   "80_From_HMI_MAN_DQ_139_4" : Bool = PLC "80_From_HMI".MAN_DQ_139_4, 1 s
   "80_From_HMI_MAN_DQ_139_5" : Bool = PLC "80_From_HMI".MAN_DQ_139_5, 1 s
   "80_From_HMI_MAN_DQ_139_6" : Bool = PLC "80_From_HMI".MAN_DQ_139_6, 1 s
   "80_From_HMI_MAN_DQ_139_7" : Bool = PLC "80_From_HMI".MAN_DQ_139_7, 1 s
   "80_From_HMI_P301_PRSNT" : Bool = PLC "80_From_HMI".P301_PRSNT, 1 s
   "80_From_HMI_P305_PRSNT" : Bool = PLC "80_From_HMI".P305_PRSNT, 1 s
   "80_From_HMI_PIT 316 delay" : Time = PLC "80_From_HMI"."PIT 316 delay", 1 s
   "80_From_HMI_PIT 359 delay" : Time = PLC "80_From_HMI"."PIT 359 delay", 1 s
   "80_From_HMI_Post Purge Time" : Time = PLC "80_From_HMI"."Post Purge Time", 1 s
   "80_From_HMI_Request_Auto" : Bool = PLC "80_From_HMI".Request_Auto, 1 s
   "80_From_HMI_Request_Manual" : Bool = PLC "80_From_HMI".Request_Manual, 1 s
   "80_From_HMI_Reset CV203 PID" : Bool = PLC "80_From_HMI"."Reset CV203 PID", 1 s
   "80_From_HMI_Reset_Alarms" : Bool = PLC "80_From_HMI".Reset_Alarms, 1 s
   "80_From_HMI_RST_AUT_SEQ" : Bool = PLC "80_From_HMI".RST_AUT_SEQ, 1 s
   "80_From_HMI_RST_LOCKOUT" : Bool = PLC "80_From_HMI".RST_LOCKOUT, 1 s
   "80_From_HMI_RUN_BTCS" : Bool = PLC "80_From_HMI".RUN_BTCS, 1 s
   "80_From_HMI_RUN_BWTS" : Bool = PLC "80_From_HMI".RUN_BWTS, 1 s
   "80_From_HMI_SAL_CNFRM" : Bool = PLC "80_From_HMI".SAL_CNFRM, 1 s
   "80_From_HMI_SAL_VALUE" : Real = PLC "80_From_HMI".SAL_VALUE, 1 s
   "80_From_HMI_Test Tank Request" : Bool = PLC "80_From_HMI"."Test Tank Request", 1 s
   "80_From_HMI_TIMER RST Supres" : Bool = PLC "80_From_HMI"."TIMER RST Supres", 1 s
   "82_To_HMI_CA Blower Reset Hours" : Bool = PLC "82_To_HMI"."CA Blower Reset Hours", 1 s
   "82_To_HMI_CA Blower Run Seconds" : Int = PLC "82_To_HMI"."CA Blower Run Seconds", 1 s
   "82_To_HMI_CA Blower Service Due" : Bool = PLC "82_To_HMI"."CA Blower Service Due", 1 s
   "82_To_HMI_CA Blower Total Run Hours" : Int = PLC "82_To_HMI"."CA Blower Total Run Hours", 1 s
   "82_To_HMI_CRNT_MODE" : Int = PLC "82_To_HMI".CRNT_MODE_IGG, 1 s
   "82_To_HMI_CRNT_MODE_GCU" : Int = PLC "82_To_HMI".CRNT_MODE_GCU, 1 s
   "82_To_HMI_E500A Fuel Pump Reset Hours" : Bool = PLC "82_To_HMI"."E500A Fuel Pump Reset Hours", 1 s
   "82_To_HMI_E500A Fuel Pump Run Hours" : Int = PLC "82_To_HMI"."E500A Fuel Pump Run Hours", 1 s
   "82_To_HMI_E500A Fuel Pump Run Minutes" : Int = PLC "82_To_HMI"."E500A Fuel Pump Run Minutes", 1 s
   "82_To_HMI_E500A Fuel Pump Run Seconds" : Int = PLC "82_To_HMI"."E500A Fuel Pump Run Seconds", 1 s
   "82_To_HMI_E500A Fuel Pump Service Due" : Bool = PLC "82_To_HMI"."E500A Fuel Pump Service Due", 1 s
   "82_To_HMI_E500A Fuel Pump Service Time Hours" : Int = PLC "82_To_HMI"."E500A Fuel Pump Service Time Hours", 1 s
   "82_To_HMI_E500A Fuel Pump Total Run Hours" : Int = PLC "82_To_HMI"."E500A Fuel Pump Total Run Hours", 1 s
   "82_To_HMI_E500B Fuel Pump Reset Hours" : Bool = PLC "82_To_HMI"."E500B Fuel Pump Reset Hours", 1 s
   "82_To_HMI_E500B Fuel Pump Run Minutes" : Int = PLC "82_To_HMI"."E500B Fuel Pump Run Minutes", 1 s
   "82_To_HMI_E500B Fuel Pump Run Seconds" : Int = PLC "82_To_HMI"."E500B Fuel Pump Run Seconds", 1 s
   "82_To_HMI_E500B Fuel Pump Service Due" : Bool = PLC "82_To_HMI"."E500B Fuel Pump Service Due", 1 s
   "82_To_HMI_E500B Fuel Pump Service Time Hours" : Int = PLC "82_To_HMI"."E500B Fuel Pump Service Time Hours", 1 s
   "82_To_HMI_E500B Fuel Pump Total Run Hours" : Int = PLC "82_To_HMI"."E500B Fuel Pump Total Run Hours", 1 s
   "82_To_HMI_E-STOP LATCHED" : Bool = PLC "82_To_HMI"."E-STOP LATCHED", 1 s
   "82_To_HMI_I&A Compressor Reset Hours" : Bool = PLC "82_To_HMI"."I&A Compressor Reset Hours", 1 s
   "82_To_HMI_I&A Compressor Service Due" : Bool = PLC "82_To_HMI"."I&A Compressor Service Due", 1 s
   "82_To_HMI_I&A Compressor Total Run Hours" : Int = PLC "82_To_HMI"."I&A Compressor Total Run Hours", 1 s
   "82_To_HMI_P301 CSW Pump Reset Hours" : Bool = PLC "82_To_HMI"."P301 CSW Pump Reset Hours", 1 s
   "82_To_HMI_P301 CSW Pump Run Days" : Int = PLC "82_To_HMI"."P301 CSW Pump Run Days", 1 s
   "82_To_HMI_P301 CSW Pump Run Hours" : Int = PLC "82_To_HMI"."P301 CSW Pump Run Hours", 1 s
   "82_To_HMI_P301 CSW Pump Run Minutes" : Int = PLC "82_To_HMI"."P301 CSW Pump Run Minutes", 1 s
   "82_To_HMI_P301 CSW Pump Run Seconds" : Int = PLC "82_To_HMI"."P301 CSW Pump Run Seconds", 1 s
   "82_To_HMI_P301 CSW Pump Service Due" : Bool = PLC "82_To_HMI"."P301 CSW Pump Service Due", 1 s
   "82_To_HMI_P301 CSW Pump Service Time Hours" : Int = PLC "82_To_HMI"."P301 CSW Pump Service Time Hours", 1 s
   "82_To_HMI_P301 CSW Pump Total Run Hours" : Int = PLC "82_To_HMI"."P301 CSW Pump Total Run Hours", 1 s
   "82_To_HMI_P305 FW Pump Reset Hours" : Bool = PLC "82_To_HMI"."P305 FW Pump Reset Hours", 1 s
   "82_To_HMI_P305 FW Pump Run Days" : Int = PLC "82_To_HMI"."P305 FW Pump Run Days", 1 s
   "82_To_HMI_P305 FW Pump Run Hours" : Int = PLC "82_To_HMI"."P305 FW Pump Run Hours", 1 s
   "84_Setpoints_D_ON" : Bool = PLC "84_Setpoints".D_ON, 1 s
   "84_Setpoints_Derive Time" : Time = PLC "84_Setpoints"."Derive Time", 1 s
   "84_Setpoints_E400_PT002_High" : Real = PLC "84_Setpoints".E400_PT002_High, 1 s
   "84_Setpoints_E400_PT002_HighHigh" : Real = PLC "84_Setpoints".E400_PT002_HighHigh, 1 s
   "84_Setpoints_E400_TT002_High" : Real = PLC "84_Setpoints".E400_TT002_High, 1 s
   "84_Setpoints_E400_TT002_HighHigh" : Real = PLC "84_Setpoints".E400_TT002_HighHigh, 1 s
   "84_Setpoints_Gain" : Real = PLC "84_Setpoints".Gain, 1 s
   "84_Setpoints_I_ON" : Bool = PLC "84_Setpoints".I_ON, 1 s
   "84_Setpoints_Integration Time" : Time = PLC "84_Setpoints"."Integration Time", 1 s
   "84_Setpoints_LIT304_InitialFill_High" : Real = PLC "84_Setpoints".LIT304_InitialFill_High, 1 s
   "84_Setpoints_LIT304_InitialFill_HighHigh" : Real = PLC "84_Setpoints".LIT304_InitialFill_HighHigh, 1 s
   "84_Setpoints_LIT304_InitialFill_Low" : Real = PLC "84_Setpoints".LIT304_InitialFill_Low, 1 s
   "84_Setpoints_LIT304_InitialFill_LowLow" : Real = PLC "84_Setpoints".LIT304_InitialFill_LowLow, 1 s
   "84_Setpoints_LIT304_InitialFill_Target" : Real = PLC "84_Setpoints".LIT304_InitialFill_Target, 1 s
   "84_Setpoints_LIT304_InitialFill_Target_Low" : Real = PLC "84_Setpoints".LIT304_InitialFill_Target_Low, 1 s
   "84_Setpoints_LIT304_Refill_High" : Real = PLC "84_Setpoints".LIT304_Refill_High, 1 s
   "84_Setpoints_LIT304_Refill_HighHigh" : Real = PLC "84_Setpoints".LIT304_Refill_HighHigh, 1 s
   "84_Setpoints_LIT304_Refill_Low" : Real = PLC "84_Setpoints".LIT304_Refill_Low, 1 s
   "84_Setpoints_LIT304_Refill_LowLow" : Real = PLC "84_Setpoints".LIT304_Refill_LowLow, 1 s
   "84_Setpoints_LIT304_Refill_Target" : Real = PLC "84_Setpoints".LIT304_Refill_Target, 1 s
   "84_Setpoints_LIT304_Refill_Target_Low" : Real = PLC "84_Setpoints".LIT304_Refill_Target_Low, 1 s
   "84_Setpoints_Max Opening" : Real = PLC "84_Setpoints"."Max Opening", 1 s
   "84_Setpoints_Min Opening" : Real = PLC "84_Setpoints"."Min Opening", 1 s
   "84_Setpoints_P_ON" : Bool = PLC "84_Setpoints".P_ON, 1 s
   "84_Setpoints_PIT113_Burner_Target" : Real = PLC "84_Setpoints".PIT113_Burner_Target, 1 s
   "84_Setpoints_PIT204_High" : Real = PLC "84_Setpoints".PIT204_High, 1 s
   "84_Setpoints_PIT204_High(1)" : Real = PLC "84_Setpoints".PIT204_High, 1 s
   "84_Setpoints_PIT204_HighHigh" : Real = PLC "84_Setpoints".PIT204_HighHigh, 1 s
   "84_Setpoints_PIT204_HighHigh(1)" : Real = PLC "84_Setpoints".PIT204_HighHigh, 1 s
   "84_Setpoints_PIT204_Low" : Real = PLC "84_Setpoints".PIT204_Low, 1 s
   "84_Setpoints_PIT204_Low(1)" : Real = PLC "84_Setpoints".PIT204_Low, 1 s
   "84_Setpoints_PIT204_LowLow" : Real = PLC "84_Setpoints".PIT204_LowLow, 1 s
   "84_Setpoints_PIT204_LowLow(1)" : Real = PLC "84_Setpoints".PIT204_LowLow, 1 s
   "84_Setpoints_PIT348_High" : Real = PLC "84_Setpoints".PIT348_High, 1 s
   "84_Setpoints_PIT348_HighHigh" : Real = PLC "84_Setpoints".PIT348_HighHigh, 1 s
   "84_Setpoints_PIT348_Low" : Real = PLC "84_Setpoints".PIT348_Low, 1 s
   "84_Setpoints_PIT348_LowLow" : Real = PLC "84_Setpoints".PIT348_LowLow, 1 s
   "84_Setpoints_PIT353_InitialFill_High" : Real = PLC "84_Setpoints".PIT353_InitialFill_High, 1 s
   "84_Setpoints_PIT353_InitialFill_HighHigh" : Real = PLC "84_Setpoints".PIT353_InitialFill_HighHigh, 1 s
   "84_Setpoints_PIT353_InitialFill_Low" : Real = PLC "84_Setpoints".PIT353_InitialFill_Low, 1 s
   "84_Setpoints_PIT353_InitialFill_LowLow" : Real = PLC "84_Setpoints".PIT353_InitialFill_LowLow, 1 s
   "84_Setpoints_PIT353_Refill_High" : Real = PLC "84_Setpoints".PIT353_Refill_High, 1 s
   "84_Setpoints_PIT353_Refill_HighHigh" : Real = PLC "84_Setpoints".PIT353_Refill_HighHigh, 1 s
   "84_Setpoints_PIT353_Refill_Low" : Real = PLC "84_Setpoints".PIT353_Refill_Low, 1 s
   "84_Setpoints_PIT353_Refill_LowLow" : Real = PLC "84_Setpoints".PIT353_Refill_LowLow, 1 s
   "84_Setpoints_PIT358_InitialFill_High" : Real = PLC "84_Setpoints".PIT358_InitialFill_High, 1 s
   "84_Setpoints_PIT358_InitialFill_HighHigh" : Real = PLC "84_Setpoints".PIT358_InitialFill_HighHigh, 1 s
   "84_Setpoints_PIT358_InitialFill_Low" : Real = PLC "84_Setpoints".PIT358_InitialFill_Low, 1 s
   "84_Setpoints_PIT358_InitialFill_LowLow" : Real = PLC "84_Setpoints".PIT358_InitialFill_LowLow, 1 s
   "84_Setpoints_PIT358_Refill_High" : Real = PLC "84_Setpoints".PIT358_Refill_High, 1 s
   "84_Setpoints_PIT358_Refill_HighHigh" : Real = PLC "84_Setpoints".PIT358_Refill_HighHigh, 1 s
   "84_Setpoints_PIT358_Refill_Low" : Real = PLC "84_Setpoints".PIT358_Refill_Low, 1 s
   "84_Setpoints_PIT358_Refill_LowLow" : Real = PLC "84_Setpoints".PIT358_Refill_LowLow, 1 s
   "84_Setpoints_PIT416_High" : Real = PLC "84_Setpoints".PIT416_High, 1 s
   "84_Setpoints_PIT416_HighHigh" : Real = PLC "84_Setpoints".PIT416_HighHigh, 1 s
   "84_Setpoints_PIT416_Low" : Real = PLC "84_Setpoints".PIT416_Low, 1 s
   "84_Setpoints_PIT416_LowLow" : Real = PLC "84_Setpoints".PIT416_LowLow, 1 s
   "84_Setpoints_PIT416_Target" : Real = PLC "84_Setpoints".PIT416_Target, 1 s
   "84_Setpoints_TIT406_High" : Real = PLC "84_Setpoints".TIT406_High, 1 s
   "84_Setpoints_TIT406_HighHigh" : Real = PLC "84_Setpoints".TIT406_HighHigh, 1 s
   "84_Setpoints_TIT408_High" : Real = PLC "84_Setpoints".TIT408_High, 1 s
   "84_Setpoints_TIT408_HighHigh" : Real = PLC "84_Setpoints".TIT408_HighHigh, 1 s
   "86_Times_CV341_CLSD_DLY" : Time = PLC "86_Times".CV341_CLSD_DLY, 1 s
   "86_Times_CV341_MAX_TRVL_TIME" : Time = PLC "86_Times".CV341_MAX_TRVL_TIME, 1 s
   "86_Times_CV341_OPND_DLY" : Time = PLC "86_Times".CV341_OPND_DLY, 1 s
   "86_Times_CV358_CLSD_DLY" : Time = PLC "86_Times".CV358_CLSD_DLY, 1 s
   "86_Times_CV358_MAX_TRVL_TIME" : Time = PLC "86_Times".CV358_MAX_TRVL_TIME, 1 s
   "86_Times_CV401_CLSD_DLY" : Time = PLC "86_Times".CV401_CLSD_DLY, 1 s
   "86_Times_CV401_OPND_DLY" : Time = PLC "86_Times".CV401_OPND_DLY, 1 s
   "86_Times_CV405_OPND_DLY" : Time = PLC "86_Times".CV405_OPND_DLY, 1 s
   "86_Times_CV406_CLSD_DLY" : Time = PLC "86_Times".CV406_CLSD_DLY, 1 s
   "86_Times_CV406_MAX_TRVL_TIME" : Time = PLC "86_Times".CV406_MAX_TRVL_TIME, 1 s
   "86_Times_CV407_MAX_TRVL_TIME" : Time = PLC "86_Times".CV407_MAX_TRVL_TIME, 1 s
   "86_Times_CV409_MAX_TRVL_TIME" : Time = PLC "86_Times".CV409_MAX_TRVL_TIME, 1 s
   "86_Times_CV411_MAX_TRVL_TIME" : Time = PLC "86_Times".CV411_MAX_TRVL_TIME, 1 s
   "86_Times_CV441_CLSD_DLY" : Time = PLC "86_Times".CV441_CLSD_DLY, 1 s
   "86_Times_CV441_MAX_TRVL_TIME" : Time = PLC "86_Times".CV441_MAX_TRVL_TIME, 1 s
   "86_Times_CV441_OPND_DLY" : Time = PLC "86_Times".CV441_OPND_DLY, 1 s
   "86_Times_E400_RNG_DLY" : Time = PLC "86_Times".E400_RNG_DLY, 1 s
   "86_Times_E400_STOP_TIME" : Time = PLC "86_Times".E400_STOP_TIME, 1 s
   "86_Times_E400_STRTD_DLY" : Time = PLC "86_Times".E400_STRTD_DLY, 1 s
   "86_Times_GCU_FLUSH_TIME" : Time = PLC "86_Times".GCU_FLUSH_TIME, 1 s
   "86_Times_GCU_TNK_DRN_MAX_TIME" : Time = PLC "86_Times".GCU_TNK_DRN_MAX_TIME, 1 s
   "86_Times_GCU_TNK_FILL_MAX_TIME" : Time = PLC "86_Times".GCU_TNK_FILL_MAX_TIME, 1 s
   "86_Times_LIT304 Delay" : Time = PLC "86_Times"."LIT304 Delay", 1 s
   "86_Times_P301_START_DLY" : Time = PLC "86_Times".P301_START_DLY, 1 s
   "86_Times_P303_STOP_TIME" : Time = PLC "86_Times".P303_STOP_TIME, 1 s
   "86_Times_P303_STPD_DLY" : Time = PLC "86_Times".P303_STPD_DLY, 1 s
   "86_Times_P303_STRTD_DLY" : Time = PLC "86_Times".P303_STRTD_DLY, 1 s
   "86_Times_P304_STPD_DLY" : Time = PLC "86_Times".P304_STPD_DLY, 1 s
   "86_Times_P304_STRTD_DLY" : Time = PLC "86_Times".P304_STRTD_DLY, 1 s
   "86_Times_P305_STPD_DLY" : Time = PLC "86_Times".P305_STPD_DLY, 1 s
   "86_Times_P305_STRTD_DLY" : Time = PLC "86_Times".P305_STRTD_DLY, 1 s
   "86_Times_PIT353 Delay" : Time = PLC "86_Times"."PIT353 Delay", 1 s
   "86_Times_PIT402 Alarm Delay" : Time = PLC "86_Times"."PIT402 Alarm Delay", 1 s
   "86_Times_PIT402_Ramp_Seconds" : Int = PLC "86_Times".PIT402_Ramp_Seconds, 1 s
   "86_Times_PIT416 Delay" : Time = PLC "86_Times"."PIT416 Delay", 1 s
   "86_Times_PIT416_TRGT_RMP_TIME" : Real = PLC "86_Times".PIT416_TRGT_RMP_TIME, 1 s
   "86_Times_POST_FLUSH_DLY" : Time = PLC "86_Times".POST_FLUSH_DLY, 1 s
   "86_Times_PRE_CV441_OPN_DLY" : Time = PLC "86_Times".PRE_CV441_OPN_DLY, 1 s
   "86_Times_PRE_GCU_TNK_FILL_DLY" : Time = PLC "86_Times".PRE_GCU_TNK_FILL_DLY, 1 s
   "86_Times_STEP_MAX_TIME_STP_001" : Time = PLC "86_Times".STEP_MAX_TIME_STP_001, 1 s
   "86_Times_STEP_MAX_TIME_STP_005" : Time = PLC "86_Times".STEP_MAX_TIME_STP_005, 1 s
   "86_Times_STEP_MAX_TIME_STP_010" : Time = PLC "86_Times".STEP_MAX_TIME_STP_010, 1 s
   "86_Times_STEP_MAX_TIME_STP_020" : Time = PLC "86_Times".STEP_MAX_TIME_STP_020, 1 s
   "86_Times_STEP_MAX_TIME_STP_030" : Time = PLC "86_Times".STEP_MAX_TIME_STP_030, 1 s
   "86_Times_STEP_MAX_TIME_STP_040" : Time = PLC "86_Times".STEP_MAX_TIME_STP_040, 1 s
   "86_Times_STEP_MAX_TIME_STP_050" : Time = PLC "86_Times".STEP_MAX_TIME_STP_050, 1 s
   "86_Times_STEP_MAX_TIME_STP_060" : Time = PLC "86_Times".STEP_MAX_TIME_STP_060, 1 s
   "86_Times_STEP_MAX_TIME_STP_070" : Time = PLC "86_Times".STEP_MAX_TIME_STP_070, 1 s
   "86_Times_STEP_MAX_TIME_STP_080" : Time = PLC "86_Times".STEP_MAX_TIME_STP_080, 1 s
   "86_Times_STEP_MAX_TIME_STP_090" : Time = PLC "86_Times".STEP_MAX_TIME_STP_090, 1 s
   "86_Times_STEP_MAX_TIME_STP_100" : Time = PLC "86_Times".STEP_MAX_TIME_STP_100, 1 s
   "86_Times_STEP_MAX_TIME_STP_110" : Time = PLC "86_Times".STEP_MAX_TIME_STP_110, 1 s
   "86_Times_STEP_MAX_TIME_STP_120" : Time = PLC "86_Times".STEP_MAX_TIME_STP_120, 1 s
   "86_Times_STEP_MAX_TIME_STP_130" : Time = PLC "86_Times".STEP_MAX_TIME_STP_130, 1 s
   "86_Times_STEP_MAX_TIME_STP_140" : Time = PLC "86_Times".STEP_MAX_TIME_STP_140, 1 s
   "86_Times_STEP_MAX_TIME_STP_150" : Time = PLC "86_Times".STEP_MAX_TIME_STP_150, 1 s
   "86_Times_STEP_MAX_TIME_STP_160" : Time = PLC "86_Times".STEP_MAX_TIME_STP_160, 1 s
   "86_Times_STEP_MAX_TIME_STP_170" : Time = PLC "86_Times".STEP_MAX_TIME_STP_170, 1 s
   "86_Times_STEP_MAX_TIME_STP_180" : Time = PLC "86_Times".STEP_MAX_TIME_STP_180, 1 s
   "86_Times_STEP_MAX_TIME_STP_190" : Time = PLC "86_Times".STEP_MAX_TIME_STP_190, 1 s
   "86_Times_STEP_MAX_TIME_STP_200" : Time = PLC "86_Times".STEP_MAX_TIME_STP_200, 1 s
   "86_Times_STEP_MAX_TIME_STP_210" : Time = PLC "86_Times".STEP_MAX_TIME_STP_210, 1 s
   "86_Times_STEP_MAX_TIME_STP_220" : Time = PLC "86_Times".STEP_MAX_TIME_STP_220, 1 s
   "86_Times_STEP_MAX_TIME_STP_230" : Time = PLC "86_Times".STEP_MAX_TIME_STP_230, 1 s
   "86_Times_STEP_MAX_TIME_STP_240" : Time = PLC "86_Times".STEP_MAX_TIME_STP_240, 1 s
   "86_Times_STEP_MAX_TIME_STP_250" : Time = PLC "86_Times".STEP_MAX_TIME_STP_250, 1 s
   "86_Times_STEP_MAX_TIME_STP_260" : Time = PLC "86_Times".STEP_MAX_TIME_STP_260, 1 s
   "86_Times_STEP_MAX_TIME_STP_270" : Time = PLC "86_Times".STEP_MAX_TIME_STP_270, 1 s
   "86_Times_STEP_MAX_TIME_STP_280" : Time = PLC "86_Times".STEP_MAX_TIME_STP_280, 1 s
   "86_Times_STEP_MAX_TIME_STP_290" : Time = PLC "86_Times".STEP_MAX_TIME_STP_290, 1 s
   "86_Times_STEP_MAX_TIME_STP_300" : Time = PLC "86_Times".STEP_MAX_TIME_STP_300, 1 s
   "86_Times_STEP_MAX_TIME_STP_310" : Time = PLC "86_Times".STEP_MAX_TIME_STP_310, 1 s
   "86_Times_STEP_MAX_TIME_STP_320" : Time = PLC "86_Times".STEP_MAX_TIME_STP_320, 1 s
   "86_Times_STEP_MAX_TIME_STP_330" : Time = PLC "86_Times".STEP_MAX_TIME_STP_330, 1 s
   "86_Times_STEP_MAX_TIME_STP_340" : Time = PLC "86_Times".STEP_MAX_TIME_STP_340, 1 s
   "86_Times_STEP_MAX_TIME_STP_350" : Time = PLC "86_Times".STEP_MAX_TIME_STP_350, 1 s
   "86_Times_STEP_MAX_TIME_STP_360" : Time = PLC "86_Times".STEP_MAX_TIME_STP_360, 1 s
   "86_Times_STEP_MAX_TIME_STP_370" : Time = PLC "86_Times".STEP_MAX_TIME_STP_370, 1 s
   "86_Times_STEP_MAX_TIME_STP_380" : Time = PLC "86_Times".STEP_MAX_TIME_STP_380, 1 s
   "86_Times_STEP_MAX_TIME_STP_390" : Time = PLC "86_Times".STEP_MAX_TIME_STP_390, 1 s
   "86_Times_STEP_MAX_TIME_STP_400" : Time = PLC "86_Times".STEP_MAX_TIME_STP_400, 1 s
   "86_Times_STEP_MAX_TIME_STP_410" : Time = PLC "86_Times".STEP_MAX_TIME_STP_410, 1 s
   "86_Times_STEP_MAX_TIME_STP_420" : Time = PLC "86_Times".STEP_MAX_TIME_STP_420, 1 s
   "86_Times_STEP_MAX_TIME_STP_430" : Time = PLC "86_Times".STEP_MAX_TIME_STP_430, 1 s
   "86_Times_STEP_MAX_TIME_STP_440" : Time = PLC "86_Times".STEP_MAX_TIME_STP_440, 1 s
   "86_Times_STEP_MAX_TIME_STP_450" : Time = PLC "86_Times".STEP_MAX_TIME_STP_450, 1 s
   "86_Times_STEP_MAX_TIME_STP_460" : Time = PLC "86_Times".STEP_MAX_TIME_STP_460, 1 s
   "86_Times_STEP_MAX_TIME_STP_470" : Time = PLC "86_Times".STEP_MAX_TIME_STP_470, 1 s
   "86_Times_STEP_MAX_TIME_STP_480" : Time = PLC "86_Times".STEP_MAX_TIME_STP_480, 1 s
   "86_Times_STEP_MAX_TIME_STP_490" : Time = PLC "86_Times".STEP_MAX_TIME_STP_490, 1 s
   "86_Times_STEP_MAX_TIME_STP_500" : Time = PLC "86_Times".STEP_MAX_TIME_STP_500, 1 s
   "86_Times_STEP_MAX_TIME_STP_510" : Time = PLC "86_Times".STEP_MAX_TIME_STP_510, 1 s
   "86_Times_STEP_MAX_TIME_STP_520" : Time = PLC "86_Times".STEP_MAX_TIME_STP_520, 1 s
   "86_Times_STEP_MAX_TIME_STP_530" : Time = PLC "86_Times".STEP_MAX_TIME_STP_530, 1 s
   "86_Times_STEP_MAX_TIME_STP_540" : Time = PLC "86_Times".STEP_MAX_TIME_STP_540, 1 s
   "86_Times_STEP_MAX_TIME_STP_550" : Time = PLC "86_Times".STEP_MAX_TIME_STP_550, 1 s
   "86_Times_STEP_MAX_TIME_STP_560" : Time = PLC "86_Times".STEP_MAX_TIME_STP_560, 1 s
   "86_Times_STEP_MAX_TIME_STP_570" : Time = PLC "86_Times".STEP_MAX_TIME_STP_570, 1 s
   "86_Times_STEP_MAX_TIME_STP_580" : Time = PLC "86_Times".STEP_MAX_TIME_STP_580, 1 s
   "86_Times_STEP_MAX_TIME_STP_590" : Time = PLC "86_Times".STEP_MAX_TIME_STP_590, 1 s
   "86_Times_STEP_MAX_TIME_STP_600" : Time = PLC "86_Times".STEP_MAX_TIME_STP_600, 1 s
   "86_Times_STEP_MAX_TIME_STP_610" : Time = PLC "86_Times".STEP_MAX_TIME_STP_610, 1 s
   "86_Times_STEP_MAX_TIME_STP_620" : Time = PLC "86_Times".STEP_MAX_TIME_STP_620, 1 s
   "86_Times_STEP_MAX_TIME_STP_630" : Time = PLC "86_Times".STEP_MAX_TIME_STP_630, 1 s
   "86_Times_VLV_CNFG_DN_DLY" : Time = PLC "86_Times".VLV_CNFG_DN_DLY, 1 s
   "88_treatment_POP_UP" : Bool = PLC "88_treatment".POP_UP AT %DB1.DBX0.0, 1 s
      on ChangeValue: "TreatmentdDailyChecks"()
   "88_treatment_POP_UP_CNFRM" : Bool = PLC "88_treatment".POP_UP_CNFRM AT %DB1.DBX0.0, 1 s
   "Activate Tank Port 1" : Bool = PLC "504_Tank Grouping_DB2020"."TANK ACTIV 2" AT %DB1.DBW0, 1 s
   "Activate Tank Port 10" : Bool = PLC "504_Tank Grouping_DB2020"."TANK ACTIV 20" AT %DB1.DBW0, 1 s
   "Activate Tank Port 2" : Bool = PLC "504_Tank Grouping_DB2020"."TANK ACTIV 4" AT %DB1.DBW0, 1 s
   "Activate Tank Port 3" : Bool = PLC "504_Tank Grouping_DB2020"."TANK ACTIV 6" AT %DB1.DBW0, 1 s
   "Activate Tank Port 4" : Bool = PLC "504_Tank Grouping_DB2020"."TANK ACTIV 8" AT %DB1.DBW0, 1 s
   "Activate Tank Port 5" : Bool = PLC "504_Tank Grouping_DB2020"."TANK ACTIV 10" AT %DB1.DBW0, 1 s
   "Activate Tank Port 6" : Bool = PLC "504_Tank Grouping_DB2020"."TANK ACTIV 12" AT %DB1.DBW0, 1 s
   "Activate Tank Port 7" : Bool = PLC "504_Tank Grouping_DB2020"."TANK ACTIV 14" AT %DB1.DBW0, 1 s
   "Activate Tank Port 8" : Bool = PLC "504_Tank Grouping_DB2020"."TANK ACTIV 16" AT %DB1.DBW0, 1 s
   "Activate Tank Port 9" : Bool = PLC "504_Tank Grouping_DB2020"."TANK ACTIV 18" AT %DB1.DBW0, 1 s
   "Activate Tank Star 1" : Bool = PLC "504_Tank Grouping_DB2020"."TANK ACTIV 3" AT %DB1.DBW0, 1 s
   "Activate Tank Star 10" : Bool = PLC "504_Tank Grouping_DB2020"."TANK ACTIV 21" AT %DB1.DBW0, 1 s
   "Activate Tank Star 2" : Bool = PLC "504_Tank Grouping_DB2020"."TANK ACTIV 5" AT %DB1.DBW0, 1 s
   "Activate Tank Star 3" : Bool = PLC "504_Tank Grouping_DB2020"."TANK ACTIV 7" AT %DB1.DBW0, 1 s
   "Activate Tank Star 4" : Bool = PLC "504_Tank Grouping_DB2020"."TANK ACTIV 9" AT %DB1.DBW0, 1 s
   "Activate Tank Star 5" : Bool = PLC "504_Tank Grouping_DB2020"."TANK ACTIV 11" AT %DB1.DBW0, 1 s
   "Activate Tank Star 6" : Bool = PLC "504_Tank Grouping_DB2020"."TANK ACTIV 13" AT %DB1.DBW0, 1 s
   "Activate Tank Star 7" : Bool = PLC "504_Tank Grouping_DB2020"."TANK ACTIV 1" AT %DB1.DBW0, 1 s
   "Activate Tank Star 8" : Bool = PLC "504_Tank Grouping_DB2020"."TANK ACTIV 17" AT %DB1.DBW0, 1 s
   "Activate Tank Star 9" : Bool = PLC "504_Tank Grouping_DB2020"."TANK ACTIV 19" AT %DB1.DBW0, 1 s
   "Alarm beacon handling_DB_Buzzer_Timer_0_Instance_Q" : Bool = PLC "Alarm beacon handling_DB".Buzzer_Timer_0_Instance.Q, 1 s
   "Alarms_Acknowledge_IGG_ALARM_ACKNLG_1" : Word = PLC Alarms_Acknowledge.IGG_ALARM_ACKNLG_1 AT %DB67.DBW0, 1 s
   "Alarms_Acknowledge_IGG_ALARM_ACKNLG_2" : Word = PLC Alarms_Acknowledge.IGG_ALARM_ACKNLG_2 AT %DB67.DBW2, 1 s
   "Alarms_Acknowledge_IGG_ALARM_ACKNLG_3" : Word = PLC Alarms_Acknowledge.IGG_ALARM_ACKNLG_3 AT %DB67.DBW4, 1 s
   "Alarms_Acknowledge_IGG_ALARM_ACKNLG_4" : Word = PLC Alarms_Acknowledge.IGG_ALARM_ACKNLG_4 AT %DB67.DBW6, 1 s
   "AlwaysTRUE" : Bool = PLC AlwaysTRUE AT %M1.2, 1 s
   "APT BWT Level High High Switch" : Bool = PLC "APT BWT Level High High Switch" AT %I78.0, 1 s
   "APT GTT Isolation Valve Feedback - Closed" : Bool = PLC "APT GTT Isolation Valve Feedback - Closed" AT %I75.1, 1 s
   "APT GTT Isolation Valve Feedback - Opened" : Bool = PLC "APT GTT Isolation Valve Feedback - Opened" AT %I75.0, 1 s
   "APT Tank Vent Valve 1 Feedback - Closed" : Bool = PLC "APT Tank Vent Valve 1 Feedback - Closed" AT %I75.3, 1 s
   "APT Tank Vent Valve 1 Feedback - Opened" : Bool = PLC "APT Tank Vent Valve 1 Feedback - Opened" AT %I75.2, 1 s
   "APT Tank Vent Valve 2 Feedback - Closed" : Bool = PLC "APT Tank Vent Valve 2 Feedback - Closed" AT %I75.5, 1 s
   "APT Tank Vent Valve 2 Feedback - Opened" : Bool = PLC "APT Tank Vent Valve 2 Feedback - Opened" AT %I75.4, 1 s
   "Atm Oxygen Content 1 Scaled" : Real = PLC "12_AI_Data".AT_O2_01_SCALED AT %DB1.DBX0.0, 1 s
   "Atm Oxygen Content 2 Scaled" : Real = PLC "12_AI_Data".AT_O2_02_SCALED AT %DB1.DBX0.0, 1 s
   "Atmospheric Alarm" : Bool = PLC "14_DQ_Data".24K2 AT %DB1.DBX0.0, 1 s
   "Atomising Air  Valve Manual Regulator" : Int, internal
   "Ballast Water Treatment Mode Enabled" : Bool = PLC "80_From_HMI".BWT_BYPASS AT %DB1.DBX0.0, 1 s
   "BC E-Stop Healthy" : Bool = PLC "10 DI_DATA".S2_8K1_OK AT %DB1.DBX0.0, 1 s
   "BC PLC Power Healthy" : Bool = PLC "10_DI_Data".BC_PLC_PWR_OK AT %DB1.DBX0.0, 1 s
   "BC_ALARM_ACKNLG_1" : Word = PLC BC_ALARM_ACKNLG_1 AT %MW24, 1 s
   "BC_ALARM_ACKNLG_2" : Word = PLC BC_ALARM_ACKNLG_2 AT %MW26, 1 s
   "BC_ALARM_ACKNLG_3" : Word = PLC BC_ALARM_ACKNLG_3 AT %MW28, 1 s
   "BC_ALARM_ACKNLG_4" : Word = PLC BC_ALARM_ACKNLG_4 AT %MW30, 1 s
   "BC_Step_Time_001" : Time = PLC "86_Times".STEP_MAX_TIME_STP_001 AT %DB1.DBW0, 1 s
   "BC_Step_Time_005" : Time = PLC "86_Times".STEP_MAX_TIME_STP_005 AT %DB1.DBW0, 1 s
   "BC_Step_Time_010" : Time = PLC "86_Times".STEP_MAX_TIME_STP_010 AT %DB1.DBW0, 1 s
   "BC_Step_Time_020" : Time = PLC "86_Times".STEP_MAX_TIME_STP_020 AT %DB1.DBW0, 1 s
   "BC_Step_Time_030" : Time = PLC "86_Times".STEP_MAX_TIME_STP_030 AT %DB1.DBW0, 1 s
   "BC_Step_Time_040" : Time = PLC "86_Times".STEP_MAX_TIME_STP_040 AT %DB1.DBW0, 1 s
   "BC_Step_Time_050" : Time = PLC "86_Times".STEP_MAX_TIME_STP_050 AT %DB1.DBW0, 1 s
   "BC_Step_Time_060" : Time = PLC "86_Times".STEP_MAX_TIME_STP_060 AT %DB1.DBW0, 1 s
   "BC_Step_Time_070" : Time = PLC "86_Times".STEP_MAX_TIME_STP_070 AT %DB1.DBW0, 1 s
   "BC_Step_Time_080" : Time = PLC "86_Times".STEP_MAX_TIME_STP_080 AT %DB1.DBW0, 1 s
   "BC_Step_Time_090" : Time = PLC "86_Times".STEP_MAX_TIME_STP_090 AT %DB1.DBW0, 1 s
   "BC_Step_Time_100" : Time = PLC "86_Times".STEP_MAX_TIME_STP_100 AT %DB1.DBW0, 1 s
   "BC_Step_Time_110" : Time = PLC "86_Times".STEP_MAX_TIME_STP_110 AT %DB1.DBW0, 1 s
   "BC_Step_Time_120" : Time = PLC "86_Times".STEP_MAX_TIME_STP_120 AT %DB1.DBW0, 1 s
   "BC_Step_Time_130" : Time = PLC "86_Times".STEP_MAX_TIME_STP_130 AT %DB1.DBW0, 1 s
   "BC_Step_Time_140" : Time = PLC "86_Times".STEP_MAX_TIME_STP_140 AT %DB1.DBW0, 1 s
   "BC_Step_Time_150" : Time = PLC "86_Times".STEP_MAX_TIME_STP_150 AT %DB1.DBW0, 1 s
   "BC_Step_Time_160" : Time = PLC "86_Times".STEP_MAX_TIME_STP_160 AT %DB1.DBW0, 1 s
   "BC_Step_Time_170" : Time = PLC "86_Times".STEP_MAX_TIME_STP_170 AT %DB1.DBW0, 1 s
   "BC_Step_Time_180" : Time = PLC "86_Times".STEP_MAX_TIME_STP_180 AT %DB1.DBW0, 1 s
   "BC_Step_Time_190" : Time = PLC "86_Times".STEP_MAX_TIME_STP_190 AT %DB1.DBW0, 1 s
   "BC_Step_Time_200" : Time = PLC "86_Times".STEP_MAX_TIME_STP_200 AT %DB1.DBW0, 1 s
   "BC_Step_Time_210" : Time = PLC "86_Times".STEP_MAX_TIME_STP_210 AT %DB1.DBW0, 1 s
   "BC_Step_Time_220" : Time = PLC "86_Times".STEP_MAX_TIME_STP_220 AT %DB1.DBW0, 1 s
   "BC_Step_Time_230" : Time = PLC "86_Times".STEP_MAX_TIME_STP_230 AT %DB1.DBW0, 1 s
   "BC_Step_Time_240" : Time = PLC "86_Times".STEP_MAX_TIME_STP_240 AT %DB1.DBW0, 1 s
   "BC_Step_Time_250" : Time = PLC "86_Times".STEP_MAX_TIME_STP_250 AT %DB1.DBW0, 1 s
   "BC_Step_Time_260" : Time = PLC "86_Times".STEP_MAX_TIME_STP_260 AT %DB1.DBW0, 1 s
   "BC_Step_Time_270" : Time = PLC "86_Times".STEP_MAX_TIME_STP_270 AT %DB1.DBW0, 1 s
   "BC_Step_Time_280" : Time = PLC "86_Times".STEP_MAX_TIME_STP_280 AT %DB1.DBW0, 1 s
   "BC_Step_Time_290" : Time = PLC "86_Times".STEP_MAX_TIME_STP_290 AT %DB1.DBW0, 1 s
   "BC_Step_Time_300" : Time = PLC "86_Times".STEP_MAX_TIME_STP_300 AT %DB1.DBW0, 1 s
   "BC_Step_Time_310" : Time = PLC "86_Times".STEP_MAX_TIME_STP_310 AT %DB1.DBW0, 1 s
   "BC_Step_Time_320" : Time = PLC "86_Times".STEP_MAX_TIME_STP_320 AT %DB1.DBW0, 1 s
   "BC_Step_Time_330" : Time = PLC "86_Times".STEP_MAX_TIME_STP_330 AT %DB1.DBW0, 1 s
   "BC_Step_Time_340" : Time = PLC "86_Times".STEP_MAX_TIME_STP_340 AT %DB1.DBW0, 1 s
   "BC_Step_Time_350" : Time = PLC "86_Times".STEP_MAX_TIME_STP_350 AT %DB1.DBW0, 1 s
   "BC_Step_Time_360" : Time = PLC "86_Times".STEP_MAX_TIME_STP_360 AT %DB1.DBW0, 1 s
   "BC_Step_Time_370" : Time = PLC "86_Times".STEP_MAX_TIME_STP_370 AT %DB1.DBW0, 1 s
   "BC_Step_Time_380" : Time = PLC "86_Times".STEP_MAX_TIME_STP_380 AT %DB1.DBW0, 1 s
   "BC_Step_Time_390" : Time = PLC "86_Times".STEP_MAX_TIME_STP_390 AT %DB1.DBW0, 1 s
   "BC_Step_Time_400" : Time = PLC "86_Times".STEP_MAX_TIME_STP_400 AT %DB1.DBW0, 1 s
   "BC_Step_Time_410" : Time = PLC "86_Times".STEP_MAX_TIME_STP_410 AT %DB1.DBW0, 1 s
   "BC_Step_Time_420" : Time = PLC "86_Times".STEP_MAX_TIME_STP_420 AT %DB1.DBW0, 1 s
   "BC_Step_Time_430" : Time = PLC "86_Times".STEP_MAX_TIME_STP_430 AT %DB1.DBW0, 1 s
   "BC_Step_Time_440" : Time = PLC "86_Times".STEP_MAX_TIME_STP_440 AT %DB1.DBW0, 1 s
   "BC_Step_Time_450" : Time = PLC "86_Times".STEP_MAX_TIME_STP_450 AT %DB1.DBW0, 1 s
   "BC_Step_Time_460" : Time = PLC "86_Times".STEP_MAX_TIME_STP_460 AT %DB1.DBW0, 1 s
   "BC_Step_Time_470" : Time = PLC "86_Times".STEP_MAX_TIME_STP_470 AT %DB1.DBW0, 1 s
   "BC_Step_Time_480" : Time = PLC "86_Times".STEP_MAX_TIME_STP_480 AT %DB1.DBW0, 1 s
   "BC_Step_Time_490" : Time = PLC "86_Times".STEP_MAX_TIME_STP_490 AT %DB1.DBW0, 1 s
   "BC_Step_Time_500" : Time = PLC "86_Times".STEP_MAX_TIME_STP_500 AT %DB1.DBW0, 1 s
   "BC_Step_Time_510" : Time = PLC "86_Times".STEP_MAX_TIME_STP_510 AT %DB1.DBW0, 1 s
   "BC_Step_Time_520" : Time = PLC "86_Times".STEP_MAX_TIME_STP_520 AT %DB1.DBW0, 1 s
   "BC_Step_Time_530" : Time = PLC "86_Times".STEP_MAX_TIME_STP_530 AT %DB1.DBW0, 1 s
   "BC_Step_Time_540" : Time = PLC "86_Times".STEP_MAX_TIME_STP_540 AT %DB1.DBW0, 1 s
   "BC_Step_Time_550" : Time = PLC "86_Times".STEP_MAX_TIME_STP_550 AT %DB1.DBW0, 1 s
   "BC_Step_Time_560" : Time = PLC "86_Times".STEP_MAX_TIME_STP_560 AT %DB1.DBW0, 1 s
   "BC_Step_Time_570" : Time = PLC "86_Times".STEP_MAX_TIME_STP_570 AT %DB1.DBW0, 1 s
   "BC_Times_CV114 Close" : Time = PLC "86_Times".CV114_CLOSE_TIME AT %DB1.DBD0, 1 s
   "BC_Times_CV114 Open" : Time = PLC "86_Times".CV114_OPEN_TIME AT %DB1.DBX0.0, 1 s
   "BC_Times_CV124 Close" : Time = PLC "86_Times".CV124_CLOSE_TIME AT %DB1.DBD0, 1 s
   "BC_Times_CV124 Close Purge" : Time = PLC "86_Times".CV124_CLOSE_TIME_PRG AT %DB1.DBX0.0, 1 s
   "BC_Times_CV124 Open" : Time = PLC "86_Times".CV124_OPEN_TIME AT %DB1.DBX0.0, 1 s
   "BC_Times_CV127 Close Time" : Time = PLC "86_Times".CV127_CLOSED_TIME AT %DB1.DBX0.0, 1 s
   "BC_Times_CV127 Open #1" : Time = PLC "86_Times".CV127_OPEN_TIME_#1 AT %DB1.DBX0.0, 1 s
   "BC_Times_CV127 Open #2" : Time = PLC "86_Times".CV127_OPEN_TIME_#2 AT %DB1.DBX0.0, 1 s
   "BC_Times_CV206 Close" : Time = PLC "86_Times".CV206_CLOSE_TIME AT %DB1.DBX0.0, 1 s
   "BC_Times_CV206 Open" : Time = PLC "86_Times".CV206_OPEN_TIME AT %DB1.DBX0.0, 1 s
   "BC_Times_CV207 Close" : Time = PLC "86_Times".CV207_CLOSE_TIME AT %DB1.DBX0.0, 1 s
   "BC_Times_CV207 Open" : Time = PLC "86_Times".CV207_OPEN_TIME AT %DB1.DBX0.0, 1 s
   "BC_Times_CV215 Close" : Time = PLC "86_Times".CV215_CLOSE_TIME AT %DB1.DBD0, 1 s
   "BC_Times_CV215 Close Purge" : Time = PLC "86_Times".CV215_CLOSE_TIME_PRG AT %DB1.DBX0.0, 1 s
   "BC_Times_CV215 Open" : Time = PLC "86_Times".CV215_OPEN_TIME AT %DB1.DBX0.0, 1 s
   "BC_Times_CV216 Close" : Time = PLC "86_Times".CV216_CLOSE_TIME AT %DB1.DBD0, 1 s
   "BC_Times_CV216 Close Purge" : Time = PLC "86_Times".CV216_CLOSE_TIME_PRG AT %DB1.DBX0.0, 1 s
   "BC_Times_CV216 Open" : Time = PLC "86_Times".CV216_OPEN_TIME AT %DB1.DBX0.0, 1 s
   "BC_Times_CV216 Open Purge" : Time = PLC "86_Times".CV216_OPEN_TIME_PRG AT %DB1.DBX0.0, 1 s
   "BC_Times_Flame Detection Delay" : Time = PLC "86_Times".FD_DET_DELAY AT %DB1.DBD0, 1 s
   "BC_Times_Flame Detection Time" : Time = PLC "86_Times".FDU_DET_TIME AT %DB1.DBD0, 1 s
   "BC_Times_Flame Verification Time" : Time = PLC "86_Times".FD_VRFCTN_TIME AT %DB1.DBD0, 1 s
   "BC_Times_Max Ignition Seq Run Time" : Time = PLC "86_Times".MAX_IGNTN_SEQ_TIME AT %DB1.DBD0, 1 s
   "BC_Times_Max Main Burner Seq Run Time" : Time = PLC "86_Times".MAX_MAIN_BURN_SEQ_TIME AT %DB1.DBD0, 1 s
   "BC_Times_Max Pilot Burner Purge Seq Run Time" : Time = PLC "86_Times".MAX_PILOT_PURGE_SEQ_TIME AT %DB1.DBD0, 1 s
   "BC_Times_O2 Check Delay" : Time = PLC "86_Times".O2_CHECK_TIME AT %DB1.DBD0, 1 s
   "BC_Times_X001 Maximum Run Time" : Time = PLC "86_Times".X001_MAX_RUN_TIME AT %DB1.DBD0, 1 s
   "BC_Times_X001 Run Confirmation Time" : Time = PLC "86_Times".X001_RUN_CNF_TIME AT %DB1.DBD0, 1 s
   "Blower Run Days" : Int = PLC "82_To_HMI"."CA Blower Run Days", 1 s
   "Blower Run Hours" : Int = PLC "82_To_HMI"."CA Blower Run Hours", 1 s
   "Blower Run Minutes" : Int = PLC "82_To_HMI"."CA Blower Run Minutes", 1 s
   "Buzzer" : Bool = PLC "14_DQ_Data".24PF4 AT %DB1.DBX0.0, 100 ms
   "Buzzer(1)" : Bool = PLC Buzzer AT %Q1.7, 1 s
   "BWT Mode Warning" : Bool = PLC "2068_Sys_Status_Data"."Not BWT mode Warning" AT %DB1.DBX0.0, 1 s
   "BWTS IG Supply Valve Close" : Bool = PLC "10_DI_Data".CV431_CLSD AT %DB1.DBX0.0, 1 s
   "BWTS IG Supply Valve Open" : Bool = PLC "10_DI_Data".CV431_OPN AT %DB1.DBX0.0, 1 s
   "CA Blower Amps Scaled" : Real = PLC "12_AI_Data".E139_AMPS_SCALED AT %DB1.DBX0.0, 1 s
   "CA Blower Animation" : Int = PLC "82_To_HMI"."CA Blower Animation" AT %DB1.DBX0.0, 100 ms
   "CA Blower Control" : Bool = PLC "14_DQ_Data".E139_CNTRL AT %DB1.DBX0.0, 1 s
   "CA Blower On" : Bool = PLC "10_DI_Data".E139_RUNNING AT %DB1.DBX0.0, 1 s
   "CA Blower Pressure Scaled" : Real = PLC "12_AI_Data".PIT102_SCALED AT %DB1.DBX0.0, 1 s
   "CA Blower Ready" : Bool = PLC "10_DI_Data".E139_READY AT %DB1.DBX0.0, 1 s
   "CA Blower RPM Scaled" : Real = PLC "12_AI_Data".E139_RPM_SCALED AT %DB1.DBX0.0, 1 s
   "CA Blower Running" : Bool = PLC "10_DI_Data".E139_RUNNING AT %DB1.DBX0.0, 1 s
   "CA Blower Speed Control" : Real = PLC "16_AQ_Data".E139_SPEED AT %DB1.DBD0, 1 s
   "CA Pressure PIT102 Scaled" : Real = PLC "12_AI_Data".PIT102_SCALED AT %DB1.DBX0.0, 1 s
   "CA Pressure Switch (PS101) Status" : Bool = PLC "10 DI_DATA".PS101 AT %DB1.DBX0.0, 1 s
   "Cargo Blanketing IG Supply Valve Close" : Bool = PLC "10_DI_Data".CV432_CLSD AT %DB1.DBX0.0, 1 s
   "Cargo Blanketing IG Supply Valve Open" : Bool = PLC "10_DI_Data".CV432_OPN AT %DB1.DBX0.0, 1 s
   "Cargo Blanketing Mode Enabled" : Bool = PLC "80_From_HMI".CRG_BLNK_MODE AT %DB1.DBX0.0, 1 s
   "Check Instrument TS403" : Bool = PLC "10 DI_DATA".TS403_FAULT AT %DB1.DBX0.0, 1 s
   "Clock_1Hz" : Bool = PLC Clock_1Hz AT %M0.5, 500 ms
   "Cooling Sea Water Pump Shutdown" : Bool = PLC "10 DI_DATA".P301_TRIPPED AT %DB1.DBX0.0, 1 s
